   Machine[2].PneumaticFlow.PV_SetV.WarningUpperLimit := 0.0;
   Machine[2].PneumaticFlow.PV_SetV.AlarmLowerLimit := 0.0;
   Machine[2].PneumaticFlow.PV_SetV.AlarmUpperLimit := 0.0;
   Machine[2].PneumaticFlow.PV_ActV.Value := 0.0;
   Machine[2].PneumaticFlow.PV_ActV.ValueState := 16#0000;
   Machine[2].PneumaticFlow.PV_Conf_ActV.ModulNo := 0;
   Machine[2].PneumaticFlow.PV_Conf_ActV.Address := 0;
   Machine[2].PneumaticFlow.PV_Conf_ActV.OffsetSignal := 0;
   Machine[2].PneumaticFlow.PV_Conf_ActV.Multiplier := 0.0;
   Machine[2].PneumaticFlow.PV_Conf_ActV.MinValueSensor := 0.0;
   Machine[2].PneumaticFlow.PV_Conf_ActV.MaxValueSensor := 0.0;
   Machine[2].PneumaticFlow.PV_Conf_ActV.MaxSignalResolution := 0.0;
END_DATA_BLOCK

DATA_BLOCK "DB608_PV_Metering"   // DB608
TITLE = Process values of metering
{ S7_Optimized_Access := 'FALSE' }
AUTHOR : KT242
VERSION : 0.1
   VAR
      ReadWriteDeviceNo : Int := 0;
      CopyDeviceNO : Int := 0;
      Read : Bool := TRUE;
      Write : Bool := FALSE;
      Copy : Bool := FALSE;
      Metering : Array[0..12] of "UDT508_PV_Metering";
      HeatexchangerHP : Array[0..12] of "UDT910_ProcessValue";
      HeatexchangerLP : Array[0..12] of "UDT910_ProcessValue";
      Heating : Array[0..4] of Struct
         Heating : Array[1..8] of "UDT910_ProcessValue";
      END_STRUCT;
   END_VAR
BEGIN
   Metering[0].Flow.PV_SetV.Value := 0.0;
   Metering[0].Flow.PV_SetV.WarningLowerLimit := 0.0;
   Metering[0].Flow.PV_SetV.WarningUpperLimit := 0.0;
   Metering[0].Flow.PV_SetV.AlarmLowerLimit := 0.0;
   Metering[0].Flow.PV_SetV.AlarmUpperLimit := 0.0;
   Metering[0].Flow.PV_ActV.Value := 0.0;
   Metering[0].Flow.PV_ActV.ValueState := 16#0000;
   Metering[0].Flow.PV_Conf_ActV.ModulNo := 0;
   Metering[0].Flow.PV_Conf_ActV.Address := 1000;
   Metering[0].Flow.PV_Conf_ActV.OffsetSignal := 0;
   Metering[0].Flow.PV_Conf_ActV.Multiplier := 0.0;
   Metering[0].Flow.PV_Conf_ActV.MinValueSensor := 0.0;
   Metering[0].Flow.PV_Conf_ActV.MaxValueSensor := 0.0;
   Metering[0].Flow.PV_Conf_ActV.MaxSignalResolution := 0.0;
   Metering[0].Pressure.PV_SetV.Value := 0.0;
   Metering[0].Pressure.PV_SetV.WarningLowerLimit := 0.0;
   Metering[0].Pressure.PV_SetV.WarningUpperLimit := 0.0;
   Metering[0].Pressure.PV_SetV.AlarmLowerLimit := 0.0;
   Metering[0].Pressure.PV_SetV.AlarmUpperLimit := 0.0;
   Metering[0].Pressure.PV_ActV.Value := 1.6;
   Metering[0].Pressure.PV_ActV.ValueState := 16#0000;
   Metering[0].Pressure.PV_Conf_ActV.ModulNo := 1;
   Metering[0].Pressure.PV_Conf_ActV.Address := 316;
   Metering[0].Pressure.PV_Conf_ActV.OffsetSignal := 0;
   Metering[0].Pressure.PV_Conf_ActV.Multiplier := 10.0;
   Metering[0].Pressure.PV_Conf_ActV.MinValueSensor := -50.0;
   Metering[0].Pressure.PV_Conf_ActV.MaxValueSensor := 60000.0;
   Metering[0].Pressure.PV_Conf_ActV.MaxSignalResolution := 0.0;
   Metering[0].Temperature.PV_SetV.Value := 0.0;
   Metering[0].Temperature.PV_SetV.WarningLowerLimit := 0.0;
   Metering[0].Temperature.PV_SetV.WarningUpperLimit := 0.0;
   Metering[0].Temperature.PV_SetV.AlarmLowerLimit := 0.0;
   Metering[0].Temperature.PV_SetV.AlarmUpperLimit := 0.0;
   Metering[0].Temperature.PV_ActV.Value := 0.0;
   Metering[0].Temperature.PV_ActV.ValueState := 16#0000;
   Metering[0].Temperature.PV_Conf_ActV.ModulNo := 0;
   Metering[0].Temperature.PV_Conf_ActV.Address := 0;
   Metering[0].Temperature.PV_Conf_ActV.OffsetSignal := 0;
   Metering[0].Temperature.PV_Conf_ActV.Multiplier := 10.0;
   Metering[0].Temperature.PV_Conf_ActV.MinValueSensor := 1.0;
   Metering[0].Temperature.PV_Conf_ActV.MaxValueSensor := 1000.0;
   Metering[0].Temperature.PV_Conf_ActV.MaxSignalResolution := 0.0;
   Metering[0].Pre_Pressure.PV_SetV.Value := 0.0;
   Metering[0].Pre_Pressure.PV_SetV.WarningLowerLimit := 0.0;
   Metering[0].Pre_Pressure.PV_SetV.WarningUpperLimit := 0.0;
   Metering[0].Pre_Pressure.PV_SetV.AlarmLowerLimit := 0.0;
   Metering[0].Pre_Pressure.PV_SetV.AlarmUpperLimit := 0.0;
   Metering[0].Pre_Pressure.PV_ActV.Value := 0.0;
   Metering[0].Pre_Pressure.PV_ActV.ValueState := 16#0000;
   Metering[0].Pre_Pressure.PV_Conf_ActV.ModulNo := 1;
   Metering[0].Pre_Pressure.PV_Conf_ActV.Address := 0;
   Metering[0].Pre_Pressure.PV_Conf_ActV.OffsetSignal := 0;
   Metering[0].Pre_Pressure.PV_Conf_ActV.Multiplier := 10.0;
   Metering[0].Pre_Pressure.PV_Conf_ActV.MinValueSensor := -50.0;
   Metering[0].Pre_Pressure.PV_Conf_ActV.MaxValueSensor := 60000.0;
   Metering[0].Pre_Pressure.PV_Conf_ActV.MaxSignalResolution := 0.0;
   Metering[0].MixingRatio.PV_SetV.Value := 100.0;
   Metering[0].MixingRatio.PV_SetV.WarningLowerLimit := 0.0;
   Metering[0].MixingRatio.PV_SetV.WarningUpperLimit := 0.0;
   Metering[0].MixingRatio.PV_SetV.AlarmLowerLimit := 0.0;
   Metering[0].MixingRatio.PV_SetV.AlarmUpperLimit := 0.0;
   Metering[0].MixingRatio.PV_ActV.Value := 0.0;
   Metering[0].MixingRatio.PV_ActV.ValueState := 16#0000;
   Metering[0].MixingRatio.PV_Conf_ActV.ModulNo := 0;
   Metering[0].MixingRatio.PV_Conf_ActV.Address := 0;
   Metering[0].MixingRatio.PV_Conf_ActV.OffsetSignal := 0;
   Metering[0].MixingRatio.PV_Conf_ActV.Multiplier := 0.0;
   Metering[0].MixingRatio.PV_Conf_ActV.MinValueSensor := 0.0;
   Metering[0].MixingRatio.PV_Conf_ActV.MaxValueSensor := 0.0;
   Metering[0].MixingRatio.PV_Conf_ActV.MaxSignalResolution := 0.0;
   Metering[1].Flow.PV_SetV.Value := 0.0;
   Metering[1].Flow.PV_SetV.WarningLowerLimit := 0.0;
   Metering[1].Flow.PV_SetV.WarningUpperLimit := 0.0;
   Metering[1].Flow.PV_SetV.AlarmLowerLimit := 0.0;
   Metering[1].Flow.PV_SetV.AlarmUpperLimit := 0.0;
   Metering[1].Flow.PV_ActV.Value := 0.0;
   Metering[1].Flow.PV_ActV.ValueState := 16#0000;
   Metering[1].Flow.PV_Conf_ActV.ModulNo := 0;
   Metering[1].Flow.PV_Conf_ActV.Address := 1000;
   Metering[1].Flow.PV_Conf_ActV.OffsetSignal := 0;
   Metering[1].Flow.PV_Conf_ActV.Multiplier := 0.0;
   Metering[1].Flow.PV_Conf_ActV.MinValueSensor := 0.0;
   Metering[1].Flow.PV_Conf_ActV.MaxValueSensor := 0.0;
   Metering[1].Flow.PV_Conf_ActV.MaxSignalResolution := 0.0;
   Metering[1].Pressure.PV_SetV.Value := 0.0;
   Metering[1].Pressure.PV_SetV.WarningLowerLimit := 0.0;
   Metering[1].Pressure.PV_SetV.WarningUpperLimit := 0.0;
   Metering[1].Pressure.PV_SetV.AlarmLowerLimit := 0.0;
   Metering[1].Pressure.PV_SetV.AlarmUpperLimit := 0.0;
   Metering[1].Pressure.PV_ActV.Value := 1.6;
   Metering[1].Pressure.PV_ActV.ValueState := 16#0000;
   Metering[1].Pressure.PV_Conf_ActV.ModulNo := 1;
   Metering[1].Pressure.PV_Conf_ActV.Address := 316;
   Metering[1].Pressure.PV_Conf_ActV.OffsetSignal := 0;
   Metering[1].Pressure.PV_Conf_ActV.Multiplier := 10.0;
   Metering[1].Pressure.PV_Conf_ActV.MinValueSensor := -50.0;
   Metering[1].Pressure.PV_Conf_ActV.MaxValueSensor := 60000.0;
   Metering[1].Pressure.PV_Conf_ActV.MaxSignalResolution := 0.0;
   Metering[1].Temperature.PV_SetV.Value := 0.0;
   Metering[1].Temperature.PV_SetV.WarningLowerLimit := 0.0;
   Metering[1].Temperature.PV_SetV.WarningUpperLimit := 0.0;
   Metering[1].Temperature.PV_SetV.AlarmLowerLimit := 0.0;
   Metering[1].Temperature.PV_SetV.AlarmUpperLimit := 0.0;
   Metering[1].Temperature.PV_ActV.Value := 0.0;
   Metering[1].Temperature.PV_ActV.ValueState := 16#0000;
   Metering[1].Temperature.PV_Conf_ActV.ModulNo := 0;
   Metering[1].Temperature.PV_Conf_ActV.Address := 0;
   Metering[1].Temperature.PV_Conf_ActV.OffsetSignal := 0;
   Metering[1].Temperature.PV_Conf_ActV.Multiplier := 10.0;
   Metering[1].Temperature.PV_Conf_ActV.MinValueSensor := 1.0;
   Metering[1].Temperature.PV_Conf_ActV.MaxValueSensor := 1000.0;
   Metering[1].Temperature.PV_Conf_ActV.MaxSignalResolution := 0.0;
   Metering[1].Pre_Pressure.PV_SetV.Value := 0.0;
   Metering[1].Pre_Pressure.PV_SetV.WarningLowerLimit := 0.0;
   Metering[1].Pre_Pressure.PV_SetV.WarningUpperLimit := 0.0;
   Metering[1].Pre_Pressure.PV_SetV.AlarmLowerLimit := 0.0;
   Metering[1].Pre_Pressure.PV_SetV.AlarmUpperLimit := 0.0;
   Metering[1].Pre_Pressure.PV_ActV.Value := 0.0;
   Metering[1].Pre_Pressure.PV_ActV.ValueState := 16#0000;
   Metering[1].Pre_Pressure.PV_Conf_ActV.ModulNo := 1;
   Metering[1].Pre_Pressure.PV_Conf_ActV.Address := 0;
   Metering[1].Pre_Pressure.PV_Conf_ActV.OffsetSignal := 0;
   Metering[1].Pre_Pressure.PV_Conf_ActV.Multiplier := 10.0;
   Metering[1].Pre_Pressure.PV_Conf_ActV.MinValueSensor := -50.0;
   Metering[1].Pre_Pressure.PV_Conf_ActV.MaxValueSensor := 60000.0;
   Metering[1].Pre_Pressure.PV_Conf_ActV.MaxSignalResolution := 0.0;
   Metering[1].MixingRatio.PV_SetV.Value := 100.0;
   Metering[1].MixingRatio.PV_SetV.WarningLowerLimit := 0.0;
   Metering[1].MixingRatio.PV_SetV.WarningUpperLimit := 0.0;
   Metering[1].MixingRatio.PV_SetV.AlarmLowerLimit := 0.0;
   Metering[1].MixingRatio.PV_SetV.AlarmUpperLimit := 0.0;
   Metering[1].MixingRatio.PV_ActV.Value := 0.0;
   Metering[1].MixingRatio.PV_ActV.ValueState := 16#0000;
   Metering[1].MixingRatio.PV_Conf_ActV.ModulNo := 0;
   Metering[1].MixingRatio.PV_Conf_ActV.Address := 0;
   Metering[1].MixingRatio.PV_Conf_ActV.OffsetSignal := 0;
   Metering[1].MixingRatio.PV_Conf_ActV.Multiplier := 0.0;
   Metering[1].MixingRatio.PV_Conf_ActV.MinValueSensor := 0.0;
   Metering[1].MixingRatio.PV_Conf_ActV.MaxValueSensor := 0.0;
   Metering[1].MixingRatio.PV_Conf_ActV.MaxSignalResolution := 0.0;
   Metering[2].Flow.PV_SetV.Value := 0.0;
   Metering[2].Flow.PV_SetV.WarningLowerLimit := 0.0;
   Metering[2].Flow.PV_SetV.WarningUpperLimit := 0.0;
   Metering[2].Flow.PV_SetV.AlarmLowerLimit := 0.0;
   Metering[2].Flow.PV_SetV.AlarmUpperLimit := 0.0;
   Metering[2].Flow.PV_ActV.Value := 0.0;
   Metering[2].Flow.PV_ActV.ValueState := 16#0000;
   Metering[2].Flow.PV_Conf_ActV.ModulNo := 0;
   Metering[2].Flow.PV_Conf_ActV.Address := 1100;
   Metering[2].Flow.PV_Conf_ActV.OffsetSignal := 0;
   Metering[2].Flow.PV_Conf_ActV.Multiplier := 0.0;
   Metering[2].Flow.PV_Conf_ActV.MinValueSensor := 0.0;
   Metering[2].Flow.PV_Conf_ActV.MaxValueSensor := 0.0;
   Metering[2].Flow.PV_Conf_ActV.MaxSignalResolution := 0.0;
   Metering[2].Pressure.PV_SetV.Value := 0.0;
   Metering[2].Pressure.PV_SetV.WarningLowerLimit := 0.0;
   Metering[2].Pressure.PV_SetV.WarningUpperLimit := 0.0;
   Metering[2].Pressure.PV_SetV.AlarmLowerLimit := 0.0;
   Metering[2].Pressure.PV_SetV.AlarmUpperLimit := 0.0;
   Metering[2].Pressure.PV_ActV.Value := 1.3;
   Metering[2].Pressure.PV_ActV.ValueState := 16#0000;
   Metering[2].Pressure.PV_Conf_ActV.ModulNo := 1;
   Metering[2].Pressure.PV_Conf_ActV.Address := 318;
   Metering[2].Pressure.PV_Conf_ActV.OffsetSignal := 0;
   Metering[2].Pressure.PV_Conf_ActV.Multiplier := 10.0;
   Metering[2].Pressure.PV_Conf_ActV.MinValueSensor := -50.0;
   Metering[2].Pressure.PV_Conf_ActV.MaxValueSensor := 60000.0;
   Metering[2].Pressure.PV_Conf_ActV.MaxSignalResolution := 0.0;
   Metering[2].Temperature.PV_SetV.Value := 0.0;
   Metering[2].Temperature.PV_SetV.WarningLowerLimit := 0.0;
   Metering[2].Temperature.PV_SetV.WarningUpperLimit := 0.0;
   Metering[2].Temperature.PV_SetV.AlarmLowerLimit := 0.0;
   Metering[2].Temperature.PV_SetV.AlarmUpperLimit := 0.0;
   Metering[2].Temperature.PV_ActV.Value := 0.0;
   Metering[2].Temperature.PV_ActV.ValueState := 16#0000;
   Metering[2].Temperature.PV_Conf_ActV.ModulNo := 0;
   Metering[2].Temperature.PV_Conf_ActV.Address := 0;
   Metering[2].Temperature.PV_Conf_ActV.OffsetSignal := 0;
   Metering[2].Temperature.PV_Conf_ActV.Multiplier := 10.0;
   Metering[2].Temperature.PV_Conf_ActV.MinValueSensor := 1.0;
   Metering[2].Temperature.PV_Conf_ActV.MaxValueSensor := 1000.0;
   Metering[2].Temperature.PV_Conf_ActV.MaxSignalResolution := 0.0;
   Metering[2].Pre_Pressure.PV_SetV.Value := 0.0;
   Metering[2].Pre_Pressure.PV_SetV.WarningLowerLimit := 0.0;
   Metering[2].Pre_Pressure.PV_SetV.WarningUpperLimit := 0.0;
   Metering[2].Pre_Pressure.PV_SetV.AlarmLowerLimit := 0.0;
   Metering[2].Pre_Pressure.PV_SetV.AlarmUpperLimit := 0.0;
   Metering[2].Pre_Pressure.PV_ActV.Value := 0.0;
   Metering[2].Pre_Pressure.PV_ActV.ValueState := 16#0000;
   Metering[2].Pre_Pressure.PV_Conf_ActV.ModulNo := 1;
   Metering[2].Pre_Pressure.PV_Conf_ActV.Address := 0;
   Metering[2].Pre_Pressure.PV_Conf_ActV.OffsetSignal := 0;
   Metering[2].Pre_Pressure.PV_Conf_ActV.Multiplier := 10.0;
   Metering[2].Pre_Pressure.PV_Conf_ActV.MinValueSensor := -50.0;
   Metering[2].Pre_Pressure.PV_Conf_ActV.MaxValueSensor := 60000.0;
   Metering[2].Pre_Pressure.PV_Conf_ActV.MaxSignalResolution := 0.0;
   Metering[2].MixingRatio.PV_SetV.Value := 16#7FBF_FFFF;
   Metering[2].MixingRatio.PV_SetV.WarningLowerLimit := 0.0;
   Metering[2].MixingRatio.PV_SetV.WarningUpperLimit := 0.0;
   Metering[2].MixingRatio.PV_SetV.AlarmLowerLimit := 0.0;
   // 1634 more start values not shown
END_DATA_BLOCK

DATA_BLOCK "DB611_Hydraulic_State"   // DB611
TITLE = Status of maschine units and foaming cycle
{ S7_Optimized_Access := 'FALSE' }
VERSION : 0.1
   VAR
      ReadDeviceNo : Int := 1;
      ActualDeviceNo : Int := 1;
      CopyDeviceNO : Int := 0;
      Spare : Int;
      Read : Bool := FALSE;
      Write : Bool := FALSE;
      Copy : Bool := FALSE;
      "Fault Exist" : Bool;
      MH_Hydraulic : Array[0..2] of "UDT021_Hydr_State";
      S_Hydraulic : Array[0..2] of "UDT021_Hydr_State";
      NZL_Hydraulic : Array[0..2] of "UDT021_Hydr_State";
   END_VAR
BEGIN
   MH_Hydraulic[0].Switch_on_Motor := FALSE;
   MH_Hydraulic[0].MH_Hyd_OK := FALSE;
   MH_Hydraulic[0].Startup_Motor_finished := FALSE;
   MH_Hydraulic[0].Switch_Hydraulic_ON_OFF := FALSE;
   MH_Hydraulic[0].FaultLevel_1 := FALSE;
   MH_Hydraulic[0].FaultLevel_2 := FALSE;
   MH_Hydraulic[0].FaultLevel_3 := FALSE;
   MH_Hydraulic[0].Fault_Exist := FALSE;
   MH_Hydraulic[0].Spare_09 := FALSE;
   MH_Hydraulic[0].Request_from_CP := FALSE;
   MH_Hydraulic[0].Act_PressureBuildUp := FALSE;
   MH_Hydraulic[0].Act_Main := FALSE;
   MH_Hydraulic[0].Act_Star := FALSE;
   MH_Hydraulic[0].Act_Delta := FALSE;
   MH_Hydraulic[0].Act_Oilcooling := FALSE;
   MH_Hydraulic[0].Spare_16 := FALSE;
   MH_Hydraulic[0].State_Hydraulic := 0;
   MH_Hydraulic[1].Switch_on_Motor := FALSE;
   MH_Hydraulic[1].MH_Hyd_OK := FALSE;
   MH_Hydraulic[1].Startup_Motor_finished := FALSE;
   MH_Hydraulic[1].Switch_Hydraulic_ON_OFF := FALSE;
   MH_Hydraulic[1].FaultLevel_1 := FALSE;
   MH_Hydraulic[1].FaultLevel_2 := FALSE;
   MH_Hydraulic[1].FaultLevel_3 := FALSE;
   MH_Hydraulic[1].Fault_Exist := FALSE;
   MH_Hydraulic[1].Spare_09 := FALSE;
   MH_Hydraulic[1].Request_from_CP := FALSE;
   MH_Hydraulic[1].Act_PressureBuildUp := FALSE;
   MH_Hydraulic[1].Act_Main := FALSE;
   MH_Hydraulic[1].Act_Star := FALSE;
   MH_Hydraulic[1].Act_Delta := FALSE;
   MH_Hydraulic[1].Act_Oilcooling := FALSE;
   MH_Hydraulic[1].Spare_16 := FALSE;
   MH_Hydraulic[1].State_Hydraulic := 0;
   MH_Hydraulic[2].Switch_on_Motor := FALSE;
   MH_Hydraulic[2].MH_Hyd_OK := FALSE;
   MH_Hydraulic[2].Startup_Motor_finished := FALSE;
   MH_Hydraulic[2].Switch_Hydraulic_ON_OFF := FALSE;
   MH_Hydraulic[2].FaultLevel_1 := FALSE;
   MH_Hydraulic[2].FaultLevel_2 := FALSE;
   MH_Hydraulic[2].FaultLevel_3 := FALSE;
   MH_Hydraulic[2].Fault_Exist := FALSE;
   MH_Hydraulic[2].Spare_09 := FALSE;
   MH_Hydraulic[2].Request_from_CP := FALSE;
   MH_Hydraulic[2].Act_PressureBuildUp := FALSE;
   MH_Hydraulic[2].Act_Main := FALSE;
   MH_Hydraulic[2].Act_Star := FALSE;
   MH_Hydraulic[2].Act_Delta := FALSE;
   MH_Hydraulic[2].Act_Oilcooling := FALSE;
   MH_Hydraulic[2].Spare_16 := FALSE;
   MH_Hydraulic[2].State_Hydraulic := 0;
   S_Hydraulic[0].Switch_on_Motor := FALSE;
   S_Hydraulic[0].MH_Hyd_OK := FALSE;
   S_Hydraulic[0].Startup_Motor_finished := FALSE;
   S_Hydraulic[0].Switch_Hydraulic_ON_OFF := FALSE;
   S_Hydraulic[0].FaultLevel_1 := FALSE;
   S_Hydraulic[0].FaultLevel_2 := FALSE;
   S_Hydraulic[0].FaultLevel_3 := FALSE;
   S_Hydraulic[0].Fault_Exist := FALSE;
   S_Hydraulic[0].Spare_09 := FALSE;
   S_Hydraulic[0].Request_from_CP := FALSE;
   S_Hydraulic[0].Act_PressureBuildUp := FALSE;
   S_Hydraulic[0].Act_Main := FALSE;
   S_Hydraulic[0].Act_Star := FALSE;
   S_Hydraulic[0].Act_Delta := FALSE;
   S_Hydraulic[0].Act_Oilcooling := FALSE;
   S_Hydraulic[0].Spare_16 := FALSE;
   S_Hydraulic[0].State_Hydraulic := 0;
   S_Hydraulic[1].Switch_on_Motor := FALSE;
   S_Hydraulic[1].MH_Hyd_OK := FALSE;
   S_Hydraulic[1].Startup_Motor_finished := FALSE;
   S_Hydraulic[1].Switch_Hydraulic_ON_OFF := FALSE;
   S_Hydraulic[1].FaultLevel_1 := FALSE;
   S_Hydraulic[1].FaultLevel_2 := FALSE;
   S_Hydraulic[1].FaultLevel_3 := FALSE;
   S_Hydraulic[1].Fault_Exist := FALSE;
   S_Hydraulic[1].Spare_09 := FALSE;
   S_Hydraulic[1].Request_from_CP := FALSE;
   S_Hydraulic[1].Act_PressureBuildUp := FALSE;
   S_Hydraulic[1].Act_Main := FALSE;
   S_Hydraulic[1].Act_Star := FALSE;
   S_Hydraulic[1].Act_Delta := FALSE;
   S_Hydraulic[1].Act_Oilcooling := FALSE;
   S_Hydraulic[1].Spare_16 := FALSE;
   S_Hydraulic[1].State_Hydraulic := 0;
   S_Hydraulic[2].Switch_on_Motor := FALSE;
   S_Hydraulic[2].MH_Hyd_OK := FALSE;
   S_Hydraulic[2].Startup_Motor_finished := FALSE;
   S_Hydraulic[2].Switch_Hydraulic_ON_OFF := FALSE;
   S_Hydraulic[2].FaultLevel_1 := FALSE;
   S_Hydraulic[2].FaultLevel_2 := FALSE;
   S_Hydraulic[2].FaultLevel_3 := FALSE;
   S_Hydraulic[2].Fault_Exist := FALSE;
   S_Hydraulic[2].Spare_09 := FALSE;
   S_Hydraulic[2].Request_from_CP := FALSE;
   S_Hydraulic[2].Act_PressureBuildUp := FALSE;
   S_Hydraulic[2].Act_Main := FALSE;
   S_Hydraulic[2].Act_Star := FALSE;
   S_Hydraulic[2].Act_Delta := FALSE;
   S_Hydraulic[2].Act_Oilcooling := FALSE;
   S_Hydraulic[2].Spare_16 := FALSE;
   S_Hydraulic[2].State_Hydraulic := 0;
   NZL_Hydraulic[0].Switch_on_Motor := FALSE;
   NZL_Hydraulic[0].MH_Hyd_OK := FALSE;
   NZL_Hydraulic[0].Startup_Motor_finished := FALSE;
   NZL_Hydraulic[0].Switch_Hydraulic_ON_OFF := FALSE;
   NZL_Hydraulic[0].FaultLevel_1 := FALSE;
   NZL_Hydraulic[0].FaultLevel_2 := FALSE;
   NZL_Hydraulic[0].FaultLevel_3 := FALSE;
   NZL_Hydraulic[0].Fault_Exist := FALSE;
   NZL_Hydraulic[0].Spare_09 := FALSE;
   NZL_Hydraulic[0].Request_from_CP := FALSE;
   NZL_Hydraulic[0].Act_PressureBuildUp := FALSE;
   NZL_Hydraulic[0].Act_Main := FALSE;
   NZL_Hydraulic[0].Act_Star := FALSE;
   NZL_Hydraulic[0].Act_Delta := FALSE;
   NZL_Hydraulic[0].Act_Oilcooling := FALSE;
   NZL_Hydraulic[0].Spare_16 := FALSE;
   NZL_Hydraulic[0].State_Hydraulic := 0;
   NZL_Hydraulic[1].Switch_on_Motor := FALSE;
   NZL_Hydraulic[1].MH_Hyd_OK := FALSE;
   NZL_Hydraulic[1].Startup_Motor_finished := FALSE;
   NZL_Hydraulic[1].Switch_Hydraulic_ON_OFF := FALSE;
   NZL_Hydraulic[1].FaultLevel_1 := FALSE;
   NZL_Hydraulic[1].FaultLevel_2 := FALSE;
   NZL_Hydraulic[1].FaultLevel_3 := FALSE;
   NZL_Hydraulic[1].Fault_Exist := FALSE;
   NZL_Hydraulic[1].Spare_09 := FALSE;
   NZL_Hydraulic[1].Request_from_CP := FALSE;
   NZL_Hydraulic[1].Act_PressureBuildUp := FALSE;
   NZL_Hydraulic[1].Act_Main := FALSE;
   NZL_Hydraulic[1].Act_Star := FALSE;
   NZL_Hydraulic[1].Act_Delta := FALSE;
   NZL_Hydraulic[1].Act_Oilcooling := FALSE;
   NZL_Hydraulic[1].Spare_16 := FALSE;
   NZL_Hydraulic[1].State_Hydraulic := 0;
   NZL_Hydraulic[2].Switch_on_Motor := FALSE;
   NZL_Hydraulic[2].MH_Hyd_OK := FALSE;
   NZL_Hydraulic[2].Startup_Motor_finished := FALSE;
   NZL_Hydraulic[2].Switch_Hydraulic_ON_OFF := FALSE;
   NZL_Hydraulic[2].FaultLevel_1 := FALSE;
   NZL_Hydraulic[2].FaultLevel_2 := FALSE;
   NZL_Hydraulic[2].FaultLevel_3 := FALSE;
   NZL_Hydraulic[2].Fault_Exist := FALSE;
   NZL_Hydraulic[2].Spare_09 := FALSE;
   NZL_Hydraulic[2].Request_from_CP := FALSE;
   NZL_Hydraulic[2].Act_PressureBuildUp := FALSE;
   NZL_Hydraulic[2].Act_Main := FALSE;
   NZL_Hydraulic[2].Act_Star := FALSE;
   NZL_Hydraulic[2].Act_Delta := FALSE;
   NZL_Hydraulic[2].Act_Oilcooling := FALSE;
   NZL_Hydraulic[2].Spare_16 := FALSE;
   NZL_Hydraulic[2].State_Hydraulic := 0;
END_DATA_BLOCK

DATA_BLOCK "DB612_Tank_State"   // DB612
TITLE = Status of maschine units and foaming cycle
{ S7_Optimized_Access := 'FALSE' }
VERSION : 0.1
   VAR
      ReadDeviceNo : Int := 1;
      ActualDeviceNo : Int := 0;
      CopyDeviceNO : Int := 0;
      Read : Bool := FALSE;
      Write : Bool := FALSE;
      Copy : Bool := FALSE;
      FaulExist : Bool := FALSE;   // Eine Störung in der Gruppe Mischkopf ist vorhanden
      FaultExists : Array[0..12] of Bool;
      Tank : Array[0..12] of "UDT102_RefillingState";
      Agitator : Array[0..12] of "UDT100_AggitatorState";
      AgitatorBarell : Array[0..12] of "UDT100_AggitatorState";
      Vacuum : Array[0..12] of "UDT106_Vacuum_Status";
      CirculationPump : Array[0..12] of "UDT101_auxiDriveState";
      Pentan : Array[0..12] of "UDT102_Pentan";
      ControllerTankTemp : Array[0..12] of "UDT105_Controller_State";   // State of different controllers
      ControllerTankJacketHeater : Array[0..12] of "UDT105_Controller_State";   // State of different controllers
      ControllerBarellTemp : Array[0..12] of "UDT105_Controller_State";   // State of different controllers
      Spezial : Struct
         State_Refilling_Poly : Int := 0;   // 1->Refilling ON; 2->Fault Refilling; 3->Refilling requested but not on
         State_Refilling_Pentan : Int := 0;   // 1->Refilling ON; 2->Fault Refilling; 3->Refilling requested but not on
         State_Refilling_Nitrogen : Int := 0;   // 1->Refilling ON; 2->Fault Refilling; 3->Refilling requested but not on
         Switch_Poly_ON_OFF : Bool := FALSE;   // Switch refilling Poly ON/OFF (external Signal)
         Switch_Pentan_ON_OFF : Bool := FALSE;   // Switch refilling Pentan ON/OFF (external Signal)
         Switch_Nitrogen_ON_OFF : Bool := FALSE;   // Switch refilling Nitrogen ON/OFF (external Signal)
         RefillingPoly_Selected : Bool := FALSE;
         RefillingPentan_Selected : Bool := FALSE;
         FillingEnds : Bool := FALSE;
         NoStartFromScales : Bool := FALSE;   // Kein Start Signal von der Waage
         FPStartExternPoly : Bool := FALSE;
         FPStartExternIso : Bool := FALSE;
         NoSourceSelected : Bool := FALSE;
      END_STRUCT;
   END_VAR
BEGIN
   FaultExists[0] := FALSE;
   FaultExists[1] := FALSE;
   FaultExists[2] := FALSE;
   FaultExists[3] := FALSE;
   FaultExists[4] := FALSE;
   FaultExists[5] := FALSE;
   FaultExists[6] := FALSE;
   FaultExists[7] := FALSE;
   FaultExists[8] := FALSE;
   FaultExists[9] := FALSE;
   FaultExists[10] := FALSE;
   FaultExists[11] := FALSE;
   FaultExists[12] := FALSE;
   Tank[0].Value_No := 37;
   Tank[0].Fault_Exist := FALSE;
   Tank[0].FaultLevel_1 := FALSE;
   Tank[0].FaultLevel_2 := FALSE;
   Tank[0].FaultLevel_3 := FALSE;
   Tank[0].Spare_1_5 := FALSE;
   Tank[0].Spare_1_6 := FALSE;
   Tank[0].Select_refilling := TRUE;
   Tank[0].Spare_2_0 := FALSE;
   Tank[0].Spare_2_1 := FALSE;
   Tank[0].Spare_2_2 := FALSE;
   Tank[0].Ramp_MH_open := TRUE;
   Tank[0].FLT_Alarm_N2 := FALSE;
   Tank[0].Preagitation_runs := FALSE;
   Tank[0].Filling_Start := FALSE;
   Tank[0].Fillingtime_runs := FALSE;
   Tank[0].Select_Filling_with_Time := FALSE;
   Tank[0].Block_is_activ := FALSE;
   Tank[0].Max_Level := TRUE;
   Tank[0].Stop_Level_Filling := TRUE;
   Tank[0].Start_Level_Filling := FALSE;
   Tank[0].Min_Level := TRUE;
   Tank[0].Enable_Agitator := TRUE;
   Tank[0].Switch_Refilling_ON_OFF := FALSE;
   Tank[0].ButtonLeakageMonitorOFF := FALSE;
   Tank[0].PreWarning_Min_Level := FALSE;
   Tank[0].Switch_DrainTank_ON_OFF := FALSE;
   Tank[0].LevelTriptray := TRUE;
   Tank[0].Switch_Refilling_from_Barrel_ON_OFF := FALSE;
   Tank[0].Spare_5_4 := FALSE;
   Tank[0].Spare_5_5 := FALSE;
   Tank[0].Spare_5_6 := FALSE;
   Tank[0].Spare_5_7 := FALSE;
   Tank[0].State_Refilling := 0;
   Tank[1].Value_No := 35;
   Tank[1].Fault_Exist := FALSE;
   Tank[1].FaultLevel_1 := FALSE;
   Tank[1].FaultLevel_2 := FALSE;
   Tank[1].FaultLevel_3 := FALSE;
   Tank[1].Spare_1_5 := FALSE;
   Tank[1].Spare_1_6 := FALSE;
   Tank[1].Select_refilling := TRUE;
   Tank[1].Spare_2_0 := FALSE;
   Tank[1].Spare_2_1 := FALSE;
   Tank[1].Spare_2_2 := FALSE;
   Tank[1].Ramp_MH_open := TRUE;
   Tank[1].FLT_Alarm_N2 := FALSE;
   Tank[1].Preagitation_runs := FALSE;
   Tank[1].Filling_Start := FALSE;
   Tank[1].Fillingtime_runs := FALSE;
   Tank[1].Select_Filling_with_Time := FALSE;
   Tank[1].Block_is_activ := FALSE;
   Tank[1].Max_Level := TRUE;
   Tank[1].Stop_Level_Filling := TRUE;
   Tank[1].Start_Level_Filling := FALSE;
   Tank[1].Min_Level := TRUE;
   Tank[1].Enable_Agitator := TRUE;
   Tank[1].Switch_Refilling_ON_OFF := FALSE;
   Tank[1].ButtonLeakageMonitorOFF := FALSE;
   Tank[1].PreWarning_Min_Level := FALSE;
   Tank[1].Switch_DrainTank_ON_OFF := FALSE;
   Tank[1].LevelTriptray := TRUE;
   Tank[1].Switch_Refilling_from_Barrel_ON_OFF := FALSE;
   Tank[1].Spare_5_4 := FALSE;
   Tank[1].Spare_5_5 := FALSE;
   Tank[1].Spare_5_6 := FALSE;
   Tank[1].Spare_5_7 := FALSE;
   Tank[1].State_Refilling := 0;
   Tank[2].Value_No := 37;
   Tank[2].Fault_Exist := FALSE;
   Tank[2].FaultLevel_1 := FALSE;
   Tank[2].FaultLevel_2 := FALSE;
   Tank[2].FaultLevel_3 := FALSE;
   Tank[2].Spare_1_5 := FALSE;
   Tank[2].Spare_1_6 := FALSE;
   Tank[2].Select_refilling := TRUE;
   Tank[2].Spare_2_0 := FALSE;
   Tank[2].Spare_2_1 := FALSE;
   Tank[2].Spare_2_2 := FALSE;
   Tank[2].Ramp_MH_open := TRUE;
   Tank[2].FLT_Alarm_N2 := FALSE;
   Tank[2].Preagitation_runs := FALSE;
   Tank[2].Filling_Start := FALSE;
   Tank[2].Fillingtime_runs := FALSE;
   Tank[2].Select_Filling_with_Time := FALSE;
   Tank[2].Block_is_activ := FALSE;
   Tank[2].Max_Level := TRUE;
   Tank[2].Stop_Level_Filling := TRUE;
   Tank[2].Start_Level_Filling := FALSE;
   Tank[2].Min_Level := TRUE;
   Tank[2].Enable_Agitator := TRUE;
   Tank[2].Switch_Refilling_ON_OFF := FALSE;
   Tank[2].ButtonLeakageMonitorOFF := FALSE;
   Tank[2].PreWarning_Min_Level := FALSE;
   Tank[2].Switch_DrainTank_ON_OFF := FALSE;
   Tank[2].LevelTriptray := TRUE;
   Tank[2].Switch_Refilling_from_Barrel_ON_OFF := FALSE;
   Tank[2].Spare_5_4 := FALSE;
   Tank[2].Spare_5_5 := FALSE;
   Tank[2].Spare_5_6 := FALSE;
   Tank[2].Spare_5_7 := FALSE;
   Tank[2].State_Refilling := 0;
   Tank[3].Value_No := 0;
   Tank[3].Fault_Exist := FALSE;
   Tank[3].FaultLevel_1 := FALSE;
   Tank[3].FaultLevel_2 := FALSE;
   Tank[3].FaultLevel_3 := FALSE;
   Tank[3].Spare_1_5 := FALSE;
   Tank[3].Spare_1_6 := FALSE;
   Tank[3].Select_refilling := FALSE;
   Tank[3].Spare_2_0 := FALSE;
   Tank[3].Spare_2_1 := FALSE;
   Tank[3].Spare_2_2 := FALSE;
   Tank[3].Ramp_MH_open := FALSE;
   Tank[3].FLT_Alarm_N2 := FALSE;
   Tank[3].Preagitation_runs := FALSE;
   Tank[3].Filling_Start := FALSE;
   Tank[3].Fillingtime_runs := FALSE;
   Tank[3].Select_Filling_with_Time := FALSE;
   Tank[3].Block_is_activ := FALSE;
   Tank[3].Max_Level := FALSE;
   Tank[3].Stop_Level_Filling := FALSE;
   Tank[3].Start_Level_Filling := FALSE;
   Tank[3].Min_Level := FALSE;
   Tank[3].Enable_Agitator := FALSE;
   Tank[3].Switch_Refilling_ON_OFF := FALSE;
   Tank[3].ButtonLeakageMonitorOFF := FALSE;
   Tank[3].PreWarning_Min_Level := FALSE;
   Tank[3].Switch_DrainTank_ON_OFF := FALSE;
   Tank[3].LevelTriptray := FALSE;
   Tank[3].Switch_Refilling_from_Barrel_ON_OFF := FALSE;
   Tank[3].Spare_5_4 := FALSE;
   Tank[3].Spare_5_5 := FALSE;
   Tank[3].Spare_5_6 := FALSE;
   Tank[3].Spare_5_7 := FALSE;
   Tank[3].State_Refilling := 0;
   Tank[4].Value_No := 0;
   Tank[4].Fault_Exist := FALSE;
   Tank[4].FaultLevel_1 := FALSE;
   Tank[4].FaultLevel_2 := FALSE;
   Tank[4].FaultLevel_3 := FALSE;
   Tank[4].Spare_1_5 := FALSE;
   Tank[4].Spare_1_6 := FALSE;
   Tank[4].Select_refilling := FALSE;
   Tank[4].Spare_2_0 := FALSE;
   Tank[4].Spare_2_1 := FALSE;
   Tank[4].Spare_2_2 := FALSE;
   Tank[4].Ramp_MH_open := FALSE;
   Tank[4].FLT_Alarm_N2 := FALSE;
   Tank[4].Preagitation_runs := FALSE;
   Tank[4].Filling_Start := FALSE;
   Tank[4].Fillingtime_runs := FALSE;
   Tank[4].Select_Filling_with_Time := FALSE;
   Tank[4].Block_is_activ := FALSE;
   Tank[4].Max_Level := FALSE;
   Tank[4].Stop_Level_Filling := FALSE;
   Tank[4].Start_Level_Filling := FALSE;
   Tank[4].Min_Level := FALSE;
   Tank[4].Enable_Agitator := FALSE;
   Tank[4].Switch_Refilling_ON_OFF := FALSE;
   Tank[4].ButtonLeakageMonitorOFF := FALSE;
   Tank[4].PreWarning_Min_Level := FALSE;
   Tank[4].Switch_DrainTank_ON_OFF := FALSE;
   Tank[4].LevelTriptray := FALSE;
   Tank[4].Switch_Refilling_from_Barrel_ON_OFF := FALSE;
   Tank[4].Spare_5_4 := FALSE;
   Tank[4].Spare_5_5 := FALSE;
   Tank[4].Spare_5_6 := FALSE;
   Tank[4].Spare_5_7 := FALSE;
   Tank[4].State_Refilling := 0;
   Tank[5].Value_No := 0;
   Tank[5].Fault_Exist := FALSE;
   Tank[5].FaultLevel_1 := FALSE;
   Tank[5].FaultLevel_2 := FALSE;
   Tank[5].FaultLevel_3 := FALSE;
   Tank[5].Spare_1_5 := FALSE;
   Tank[5].Spare_1_6 := FALSE;
   Tank[5].Select_refilling := FALSE;
   Tank[5].Spare_2_0 := FALSE;
   Tank[5].Spare_2_1 := FALSE;
   Tank[5].Spare_2_2 := FALSE;
   Tank[5].Ramp_MH_open := FALSE;
   Tank[5].FLT_Alarm_N2 := FALSE;
   Tank[5].Preagitation_runs := FALSE;
   Tank[5].Filling_Start := FALSE;
   Tank[5].Fillingtime_runs := FALSE;
   Tank[5].Select_Filling_with_Time := FALSE;
   // 2231 more start values not shown
END_DATA_BLOCK

DATA_BLOCK "DB613_Komponent_State"   // DB613
TITLE = Status of maschine units and foaming cycle
{ S7_Optimized_Access := 'FALSE' }
VERSION : 0.1
   VAR
      ReadDeviceNo : Int := 1;
      ActualDeviceNo : Int;
      CopyDeviceNO : Int;
      Read : Bool;
      Write : Bool;
      Copy : Bool;
      FaulExist : Bool;   // Eine Störung in der Gruppe Mischkopf ist vorhanden
      EdgeFilter : Array[0..12] of "UDT100_EdgeFilter";
      FeedPump : Array[0..12] of "UDT100_FeedingPump";
      MeteringPump : Array[0..12] of "UDT053_Pump";
      Cylinder : Array[0..12] of "UDT062_Cylinder";
      FlowPumpMin : Array[0..12] of Real;   // Minimum flow of pump g/sec
      FlowPumpMax : Array[0..12] of Real;   // Maximum flow of pump g/sec
      FlowPump : Array[0..12] of Real;   // Set values of flow rates metering units
      FlowPumpQPB : Array[0..12] of Real;   // Set values of flow rates metering units to start quick pressure build up
      PressurePumpQPB : Array[0..12] of Real;   // Set values pressure metering units to start quick pressure build up
      FlowPumpPContr : Array[0..12] of Real;   // Set values of flow rates metering units depending on mould pressure
      AbortComponent : Array[0..12] of "UDT108_AbortComponent";
      ServoECylinder : Array[0..12] of "UDT254_ServoECylinder";
      GroupStatus : Array[0..12] of Struct
         ColorTankFlow : Byte;
         FaultExist : Bool;
      END_STRUCT;
      HeatexchangerHP : Array[0..12] of "UDT106_ControllerHeatExchanger";
      HeatexchangerLP : Array[0..12] of "UDT106_ControllerHeatExchanger";
      FeedingPumpControler : Array[0..12] of Struct
         Status : Array[0..125] of Byte;
      END_STRUCT;
      Heating : Array[0..12] of Struct   // State of different controllers
         Heating : Array[1..8] of "UDT105_ControllerHeating";
      END_STRUCT;
   END_VAR
BEGIN
END_DATA_BLOCK

DATA_BLOCK "DB614_MH_State"   // DB614
TITLE = Status of maschine units and foaming cycle
{ S7_Optimized_Access := 'FALSE' }
VERSION : 0.1
   VAR
      ReadDeviceNo : Int := 1;
      ActualDeviceNo : Int;
      CopyDeviceNO : Int;
      Spare : Int;
      Read : Bool;
      Write : Bool;
      Copy : Bool;
      InUse : Bool;
      ImpRead : Bool;
      FaulExist : Bool;   // Eine Störung in der Gruppe Mischkopf ist vorhanden
      MH_Connection : Array[0..16] of "UDT1003_MH_Connection_State";
      MH_Status : Array[0..16] of "UDT1004_MH_Status";
      MH_CleaningPiston : Array[0..16] of "UDT071_CPiston_State";
      MH_Lock : Array[0..16] of "UDT046_MH_Lock";
      InertingMH : Array[0..16] of "UDT124_Inerting";
      ShotAdjustMH : Array[0..16] of "UDT316_StateShotAdjust";
   END_VAR
BEGIN
END_DATA_BLOCK

